   // hmiStns[3].wip[11].pnCode[4] := 1000;
   // hmiStns[3].wip[11].pnCode[5] := 1000;
   // hmiStns[3].wip[11].pnCode[6] := 1000;
   // hmiStns[3].wip[11].pnCode[7] := 1000;
   // hmiStns[3].wip[12].pnCode[0] := 1000;
   // hmiStns[3].wip[12].pnCode[1] := 1000;
   // hmiStns[3].wip[12].pnCode[2] := 1000;
   // hmiStns[3].wip[12].pnCode[3] := 1000;
   // hmiStns[3].wip[12].pnCode[4] := 1000;
   // hmiStns[3].wip[12].pnCode[5] := 1000;
   // hmiStns[3].wip[12].pnCode[6] := 1000;
   // hmiStns[3].wip[12].pnCode[7] := 1000;
   // hmiStns[3].wip[13].pnCode[0] := 1000;
   // hmiStns[3].wip[13].pnCode[1] := 1000;
   // hmiStns[3].wip[13].pnCode[2] := 1000;
   // hmiStns[3].wip[13].pnCode[3] := 1000;
   // hmiStns[3].wip[13].pnCode[4] := 1000;
   // hmiStns[3].wip[13].pnCode[5] := 1000;
   // hmiStns[3].wip[13].pnCode[6] := 1000;
   // hmiStns[3].wip[13].pnCode[7] := 1000;
   // hmiStns[3].wip[14].pnCode[0] := 1000;
   // hmiStns[3].wip[14].pnCode[1] := 1000;
   // hmiStns[3].wip[14].pnCode[2] := 1000;
   // hmiStns[3].wip[14].pnCode[3] := 1000;
   // hmiStns[3].wip[14].pnCode[4] := 1000;
   // hmiStns[3].wip[14].pnCode[5] := 1000;
   // hmiStns[3].wip[14].pnCode[6] := 1000;
   // hmiStns[3].wip[14].pnCode[7] := 1000;
   // hmiStns[3].wip[15].pnCode[0] := 1000;
   // hmiStns[3].wip[15].pnCode[1] := 1000;
   // hmiStns[3].wip[15].pnCode[2] := 1000;
   // hmiStns[3].wip[15].pnCode[3] := 1000;
   // hmiStns[3].wip[15].pnCode[4] := 1000;
   // hmiStns[3].wip[15].pnCode[5] := 1000;
   // hmiStns[3].wip[15].pnCode[6] := 1000;
   // hmiStns[3].wip[15].pnCode[7] := 1000;
   // hmiStns[3].wip[16].pnCode[0] := 1000;
   // hmiStns[3].wip[16].pnCode[1] := 1000;
   // hmiStns[3].wip[16].pnCode[2] := 1000;
   // hmiStns[3].wip[16].pnCode[3] := 1000;
   // hmiStns[3].wip[16].pnCode[4] := 1000;
   // hmiStns[3].wip[16].pnCode[5] := 1000;
   // hmiStns[3].wip[16].pnCode[6] := 1000;
   // hmiStns[3].wip[16].pnCode[7] := 1000;
   // hmiStns[3].wip[17].pnCode[0] := 1000;
   // hmiStns[3].wip[17].pnCode[1] := 1000;
   // hmiStns[3].wip[17].pnCode[2] := 1000;
   // hmiStns[3].wip[17].pnCode[3] := 1000;
   // hmiStns[3].wip[17].pnCode[4] := 1000;
   // hmiStns[3].wip[17].pnCode[5] := 1000;
   // hmiStns[3].wip[17].pnCode[6] := 1000;
   // hmiStns[3].wip[17].pnCode[7] := 1000;
   // hmiStns[3].wip[18].pnCode[0] := 1000;
   // hmiStns[3].wip[18].pnCode[1] := 1000;
   // hmiStns[3].wip[18].pnCode[2] := 1000;
   // hmiStns[3].wip[18].pnCode[3] := 1000;
   // hmiStns[3].wip[18].pnCode[4] := 1000;
   // hmiStns[3].wip[18].pnCode[5] := 1000;
   // hmiStns[3].wip[18].pnCode[6] := 1000;
   // hmiStns[3].wip[18].pnCode[7] := 1000;
   // hmiStns[3].wip[19].pnCode[0] := 1000;
   // hmiStns[3].wip[19].pnCode[1] := 1000;
   // hmiStns[3].wip[19].pnCode[2] := 1000;
   // hmiStns[3].wip[19].pnCode[3] := 1000;
   // hmiStns[3].wip[19].pnCode[4] := 1000;
   // hmiStns[3].wip[19].pnCode[5] := 1000;
   // hmiStns[3].wip[19].pnCode[6] := 1000;
   // hmiStns[3].wip[19].pnCode[7] := 1000;
   // hmiStns[3].wip[20].pnCode[0] := 1000;
   // hmiStns[3].wip[20].pnCode[1] := 1000;
   // hmiStns[3].wip[20].pnCode[2] := 1000;
   // hmiStns[3].wip[20].pnCode[3] := 1000;
   // hmiStns[3].wip[20].pnCode[4] := 1000;
   // hmiStns[3].wip[20].pnCode[5] := 1000;
   // hmiStns[3].wip[20].pnCode[6] := 1000;
   // hmiStns[3].wip[20].pnCode[7] := 1000;
   // hmiStns[3].wip[21].pnCode[0] := 1000;
   // hmiStns[3].wip[21].pnCode[1] := 1000;
   // hmiStns[3].wip[21].pnCode[2] := 1000;
   // hmiStns[3].wip[21].pnCode[3] := 1000;
   // hmiStns[3].wip[21].pnCode[4] := 1000;
   // hmiStns[3].wip[21].pnCode[5] := 1000;
   // hmiStns[3].wip[21].pnCode[6] := 1000;
   // hmiStns[3].wip[21].pnCode[7] := 1000;
   // hmiStns[3].wip[22].pnCode[0] := 1000;
   // hmiStns[3].wip[22].pnCode[1] := 1000;
   // hmiStns[3].wip[22].pnCode[2] := 1000;
   // hmiStns[3].wip[22].pnCode[3] := 1000;
   // hmiStns[3].wip[22].pnCode[4] := 1000;
   // hmiStns[3].wip[22].pnCode[5] := 1000;
   // hmiStns[3].wip[22].pnCode[6] := 1000;
   // hmiStns[3].wip[22].pnCode[7] := 1000;
   // hmiStns[3].wip[23].pnCode[0] := 1000;
   // hmiStns[3].wip[23].pnCode[1] := 1000;
   // hmiStns[3].wip[23].pnCode[2] := 1000;
   // hmiStns[3].wip[23].pnCode[3] := 1000;
   // hmiStns[3].wip[23].pnCode[4] := 1000;
   // hmiStns[3].wip[23].pnCode[5] := 1000;
   // hmiStns[3].wip[23].pnCode[6] := 1000;
   // hmiStns[3].wip[23].pnCode[7] := 1000;
   // hmiStns[3].wip[24].pnCode[0] := 1000;
   // hmiStns[3].wip[24].pnCode[1] := 1000;
   // hmiStns[3].wip[24].pnCode[2] := 1000;
   // hmiStns[3].wip[24].pnCode[3] := 1000;
   // hmiStns[3].wip[24].pnCode[4] := 1000;
   // hmiStns[3].wip[24].pnCode[5] := 1000;
   // hmiStns[3].wip[24].pnCode[6] := 1000;
   // hmiStns[3].wip[24].pnCode[7] := 1000;
   // hmiStns[3].wip[25].pnCode[0] := 1000;
   // hmiStns[3].wip[25].pnCode[1] := 1000;
   // hmiStns[3].wip[25].pnCode[2] := 1000;
   // hmiStns[3].wip[25].pnCode[3] := 1000;
   // hmiStns[3].wip[25].pnCode[4] := 1000;
   // hmiStns[3].wip[25].pnCode[5] := 1000;
   // hmiStns[3].wip[25].pnCode[6] := 1000;
   // hmiStns[3].wip[25].pnCode[7] := 1000;
   // hmiStns[3].wip[26].pnCode[0] := 1000;
   // hmiStns[3].wip[26].pnCode[1] := 1000;
   // hmiStns[3].wip[26].pnCode[2] := 1000;
   // hmiStns[3].wip[26].pnCode[3] := 1000;
   // hmiStns[3].wip[26].pnCode[4] := 1000;
   // hmiStns[3].wip[26].pnCode[5] := 1000;
   // hmiStns[3].wip[26].pnCode[6] := 1000;
   // hmiStns[3].wip[26].pnCode[7] := 1000;
   // hmiStns[3].wip[27].pnCode[0] := 1000;
   // hmiStns[3].wip[27].pnCode[1] := 1000;
   // hmiStns[3].wip[27].pnCode[2] := 1000;
   // hmiStns[3].wip[27].pnCode[3] := 1000;
   // hmiStns[3].wip[27].pnCode[4] := 1000;
   // hmiStns[3].wip[27].pnCode[5] := 1000;
   // hmiStns[3].wip[27].pnCode[6] := 1000;
   // hmiStns[3].wip[27].pnCode[7] := 1000;
   // hmiStns[3].wip[28].pnCode[0] := 1000;
   // hmiStns[3].wip[28].pnCode[1] := 1000;
   // hmiStns[3].wip[28].pnCode[2] := 1000;
   // hmiStns[3].wip[28].pnCode[3] := 1000;
   // hmiStns[3].wip[28].pnCode[4] := 1000;
   // hmiStns[3].wip[28].pnCode[5] := 1000;
   // hmiStns[3].wip[28].pnCode[6] := 1000;
   // hmiStns[3].wip[28].pnCode[7] := 1000;
   // hmiStns[3].wip[29].pnCode[0] := 1000;
   // hmiStns[3].wip[29].pnCode[1] := 1000;
   // hmiStns[3].wip[29].pnCode[2] := 1000;
   // hmiStns[3].wip[29].pnCode[3] := 1000;
   // hmiStns[3].wip[29].pnCode[4] := 1000;
   // hmiStns[3].wip[29].pnCode[5] := 1000;
   // hmiStns[3].wip[29].pnCode[6] := 1000;
   // hmiStns[3].wip[29].pnCode[7] := 1000;
   // hmiStns[3].wip[30].pnCode[0] := 1000;
   // hmiStns[3].wip[30].pnCode[1] := 1000;
   // hmiStns[3].wip[30].pnCode[2] := 1000;
   // hmiStns[3].wip[30].pnCode[3] := 1000;
   // hmiStns[3].wip[30].pnCode[4] := 1000;
   // hmiStns[3].wip[30].pnCode[5] := 1000;
   // hmiStns[3].wip[30].pnCode[6] := 1000;
   // hmiStns[3].wip[30].pnCode[7] := 1000;
   // hmiStns[3].wip[31].pnCode[0] := 1000;
   // hmiStns[3].wip[31].pnCode[1] := 1000;
   // hmiStns[3].wip[31].pnCode[2] := 1000;
   // hmiStns[3].wip[31].pnCode[3] := 1000;
   // hmiStns[3].wip[31].pnCode[4] := 1000;
   // hmiStns[3].wip[31].pnCode[5] := 1000;
   // hmiStns[3].wip[31].pnCode[6] := 1000;
   // hmiStns[3].wip[31].pnCode[7] := 1000;
   // hmiStns[3].wip[32].pnCode[0] := 1000;
   // hmiStns[3].wip[32].pnCode[1] := 1000;
   // hmiStns[3].wip[32].pnCode[2] := 1000;
   // hmiStns[3].wip[32].pnCode[3] := 1000;
   // hmiStns[3].wip[32].pnCode[4] := 1000;
   // hmiStns[3].wip[32].pnCode[5] := 1000;
   // hmiStns[3].wip[32].pnCode[6] := 1000;
   // hmiStns[3].wip[32].pnCode[7] := 1000;
   // hmiStns[3].wip[33].pnCode[0] := 1000;
   // hmiStns[3].wip[33].pnCode[1] := 1000;
   // hmiStns[3].wip[33].pnCode[2] := 1000;
   // hmiStns[3].wip[33].pnCode[3] := 1000;
   // hmiStns[3].wip[33].pnCode[4] := 1000;
   // hmiStns[3].wip[33].pnCode[5] := 1000;
   // hmiStns[3].wip[33].pnCode[6] := 1000;
   // hmiStns[3].wip[33].pnCode[7] := 1000;
   // hmiStns[3].wip[34].pnCode[0] := 1000;
   // hmiStns[3].wip[34].pnCode[1] := 1000;
   // hmiStns[3].wip[34].pnCode[2] := 1000;
   // hmiStns[3].wip[34].pnCode[3] := 1000;
   // hmiStns[3].wip[34].pnCode[4] := 1000;
   // hmiStns[3].wip[34].pnCode[5] := 1000;
   // hmiStns[3].wip[34].pnCode[6] := 1000;
   // hmiStns[3].wip[34].pnCode[7] := 1000;
   // hmiStns[3].wip[35].pnCode[0] := 1000;
   // hmiStns[3].wip[35].pnCode[1] := 1000;
   // hmiStns[3].wip[35].pnCode[2] := 1000;
   // hmiStns[3].wip[35].pnCode[3] := 1000;
   // hmiStns[3].wip[35].pnCode[4] := 1000;
   // hmiStns[3].wip[35].pnCode[5] := 1000;
   // hmiStns[3].wip[35].pnCode[6] := 1000;
   // hmiStns[3].wip[35].pnCode[7] := 1000;
   // hmiStns[3].wip[36].pnCode[0] := 1000;
   // hmiStns[3].wip[36].pnCode[1] := 1000;
   // hmiStns[3].wip[36].pnCode[2] := 1000;
   // hmiStns[3].wip[36].pnCode[3] := 1000;
   // hmiStns[3].wip[36].pnCode[4] := 1000;
   // hmiStns[3].wip[36].pnCode[5] := 1000;
   // hmiStns[3].wip[36].pnCode[6] := 1000;
   // hmiStns[3].wip[36].pnCode[7] := 1000;
   // hmiStns[3].wip[37].pnCode[0] := 1000;
   // hmiStns[3].wip[37].pnCode[1] := 1000;
   // hmiStns[3].wip[37].pnCode[2] := 1000;
   // hmiStns[3].wip[37].pnCode[3] := 1000;
   // hmiStns[3].wip[37].pnCode[4] := 1000;
   // hmiStns[3].wip[37].pnCode[5] := 1000;
   // hmiStns[3].wip[37].pnCode[6] := 1000;
   // hmiStns[3].wip[37].pnCode[7] := 1000;
   // hmiStns[3].wip[38].pnCode[0] := 1000;
   // hmiStns[3].wip[38].pnCode[1] := 1000;
   // hmiStns[3].wip[38].pnCode[2] := 1000;
   // hmiStns[3].wip[38].pnCode[3] := 1000;
   // hmiStns[3].wip[38].pnCode[4] := 1000;
   // hmiStns[3].wip[38].pnCode[5] := 1000;
   // hmiStns[3].wip[38].pnCode[6] := 1000;
   // hmiStns[3].wip[38].pnCode[7] := 1000;
   // hmiStns[3].wip[39].pnCode[0] := 1000;
   // hmiStns[3].wip[39].pnCode[1] := 1000;
   // hmiStns[3].wip[39].pnCode[2] := 1000;
   // hmiStns[3].wip[39].pnCode[3] := 1000;
   // hmiStns[3].wip[39].pnCode[4] := 1000;
   // hmiStns[3].wip[39].pnCode[5] := 1000;
   // hmiStns[3].wip[39].pnCode[6] := 1000;
   // hmiStns[3].wip[39].pnCode[7] := 1000;
   // hmiStns[3].wip[40].pnCode[0] := 1000;
   // hmiStns[3].wip[40].pnCode[1] := 1000;
   // hmiStns[3].wip[40].pnCode[2] := 1000;
   // hmiStns[3].wip[40].pnCode[3] := 1000;
   // hmiStns[3].wip[40].pnCode[4] := 1000;
   // hmiStns[3].wip[40].pnCode[5] := 1000;
   // hmiStns[3].wip[40].pnCode[6] := 1000;
   // hmiStns[3].wip[40].pnCode[7] := 1000;
   // hmiStns[3].wip[41].pnCode[0] := 1000;
   // hmiStns[3].wip[41].pnCode[1] := 1000;
   // hmiStns[3].wip[41].pnCode[2] := 1000;
   // hmiStns[3].wip[41].pnCode[3] := 1000;
   // hmiStns[3].wip[41].pnCode[4] := 1000;
   // hmiStns[3].wip[41].pnCode[5] := 1000;
   // hmiStns[3].wip[41].pnCode[6] := 1000;
   // hmiStns[3].wip[41].pnCode[7] := 1000;
   // hmiStns[3].wip[42].pnCode[0] := 1000;
   // hmiStns[3].wip[42].pnCode[1] := 1000;
   // hmiStns[3].wip[42].pnCode[2] := 1000;
   // hmiStns[3].wip[42].pnCode[3] := 1000;
   // hmiStns[3].wip[42].pnCode[4] := 1000;
   // hmiStns[3].wip[42].pnCode[5] := 1000;
   // hmiStns[3].wip[42].pnCode[6] := 1000;
   // hmiStns[3].wip[42].pnCode[7] := 1000;
   // hmiStns[3].wip[43].pnCode[0] := 1000;
   // hmiStns[3].wip[43].pnCode[1] := 1000;
   // hmiStns[3].wip[43].pnCode[2] := 1000;
   // hmiStns[3].wip[43].pnCode[3] := 1000;
   // hmiStns[3].wip[43].pnCode[4] := 1000;
   // hmiStns[3].wip[43].pnCode[5] := 1000;
   // hmiStns[3].wip[43].pnCode[6] := 1000;
   // hmiStns[3].wip[43].pnCode[7] := 1000;
   // hmiStns[3].wip[44].pnCode[0] := 1000;
   // hmiStns[3].wip[44].pnCode[1] := 1000;
   // hmiStns[3].wip[44].pnCode[2] := 1000;
   // hmiStns[3].wip[44].pnCode[3] := 1000;
   // hmiStns[3].wip[44].pnCode[4] := 1000;
   // hmiStns[3].wip[44].pnCode[5] := 1000;
   // hmiStns[3].wip[44].pnCode[6] := 1000;
   // hmiStns[3].wip[44].pnCode[7] := 1000;
   // hmiStns[3].wip[45].pnCode[0] := 1000;
   // hmiStns[3].wip[45].pnCode[1] := 1000;
   // hmiStns[3].wip[45].pnCode[2] := 1000;
   // hmiStns[3].wip[45].pnCode[3] := 1000;
   // hmiStns[3].wip[45].pnCode[4] := 1000;
   // hmiStns[3].wip[45].pnCode[5] := 1000;
   // hmiStns[3].wip[45].pnCode[6] := 1000;
   // hmiStns[3].wip[45].pnCode[7] := 1000;
   // hmiStns[3].wip[46].pnCode[0] := 1000;
   // hmiStns[3].wip[46].pnCode[1] := 1000;
   // hmiStns[3].wip[46].pnCode[2] := 1000;
   // hmiStns[3].wip[46].pnCode[3] := 1000;
   // hmiStns[3].wip[46].pnCode[4] := 1000;
   // hmiStns[3].wip[46].pnCode[5] := 1000;
   // hmiStns[3].wip[46].pnCode[6] := 1000;
   // hmiStns[3].wip[46].pnCode[7] := 1000;
   // hmiStns[3].wip[47].pnCode[0] := 1000;
   // hmiStns[3].wip[47].pnCode[1] := 1000;
   // hmiStns[3].wip[47].pnCode[2] := 1000;
   // hmiStns[3].wip[47].pnCode[3] := 1000;
   // hmiStns[3].wip[47].pnCode[4] := 1000;
   // hmiStns[3].wip[47].pnCode[5] := 1000;
   // hmiStns[3].wip[47].pnCode[6] := 1000;
   // hmiStns[3].wip[47].pnCode[7] := 1000;
   // hmiStns[3].wip[48].pnCode[0] := 1000;
   // hmiStns[3].wip[48].pnCode[1] := 1000;
   // hmiStns[3].wip[48].pnCode[2] := 1000;
   // hmiStns[3].wip[48].pnCode[3] := 1000;
   // hmiStns[3].wip[48].pnCode[4] := 1000;
   // hmiStns[3].wip[48].pnCode[5] := 1000;
   // hmiStns[3].wip[48].pnCode[6] := 1000;
   // hmiStns[3].wip[48].pnCode[7] := 1000;
   // hmiStns[3].wip[49].pnCode[0] := 1000;
   // hmiStns[3].wip[49].pnCode[1] := 1000;
   // hmiStns[3].wip[49].pnCode[2] := 1000;
   // hmiStns[3].wip[49].pnCode[3] := 1000;
   // hmiStns[3].wip[49].pnCode[4] := 1000;
   // hmiStns[3].wip[49].pnCode[5] := 1000;
   // hmiStns[3].wip[49].pnCode[6] := 1000;
   // hmiStns[3].wip[49].pnCode[7] := 1000;
   // hmiStns[4].pStn := 29;
   // hmiStns[4].wip[0].pnCode[0] := 1000;
   // hmiStns[4].wip[0].pnCode[1] := 244000;
   // hmiStns[4].wip[0].pnCode[2] := 1000;
   // hmiStns[4].wip[0].pnCode[3] := 4000;
   // hmiStns[4].wip[0].pnCode[4] := 1000;
   // hmiStns[4].wip[0].pnCode[5] := 1000;
   // hmiStns[4].wip[0].pnCode[6] := 2000;
   // hmiStns[4].wip[0].pnCode[7] := 3000;
   // hmiStns[4].wip[1].pnCode[0] := 1000;
   // hmiStns[4].wip[1].pnCode[1] := 244000;
   // hmiStns[4].wip[1].pnCode[2] := 6000;
   // hmiStns[4].wip[1].pnCode[3] := 10000;
   // hmiStns[4].wip[1].pnCode[4] := 1000;
   // hmiStns[4].wip[1].pnCode[5] := 7000;
   // hmiStns[4].wip[1].pnCode[6] := 5000;
   // hmiStns[4].wip[1].pnCode[7] := 11000;
   // hmiStns[4].wip[2].pnCode[0] := 1000;
   // hmiStns[4].wip[2].pnCode[1] := 244000;
   // hmiStns[4].wip[2].pnCode[2] := 8000;
   // hmiStns[4].wip[2].pnCode[3] := 10000;
   // hmiStns[4].wip[2].pnCode[4] := 1000;
   // hmiStns[4].wip[2].pnCode[5] := 9000;
   // hmiStns[4].wip[2].pnCode[6] := 5000;
   // hmiStns[4].wip[2].pnCode[7] := 11000;
   // hmiStns[4].wip[3].pnCode[0] := 1000;
   // hmiStns[4].wip[3].pnCode[1] := 1000;
   // hmiStns[4].wip[3].pnCode[2] := 1000;
   // hmiStns[4].wip[3].pnCode[3] := 1000;
   // hmiStns[4].wip[3].pnCode[4] := 1000;
   // hmiStns[4].wip[3].pnCode[5] := 1000;
   // hmiStns[4].wip[3].pnCode[6] := 1000;
   // hmiStns[4].wip[3].pnCode[7] := 1000;
   // hmiStns[4].wip[4].pnCode[0] := 1000;
   // hmiStns[4].wip[4].pnCode[1] := 1000;
   // hmiStns[4].wip[4].pnCode[2] := 1000;
   // hmiStns[4].wip[4].pnCode[3] := 1000;
   // hmiStns[4].wip[4].pnCode[4] := 1000;
   // hmiStns[4].wip[4].pnCode[5] := 1000;
   // hmiStns[4].wip[4].pnCode[6] := 1000;
   // hmiStns[4].wip[4].pnCode[7] := 1000;
   // hmiStns[4].wip[5].pnCode[0] := 1000;
   // hmiStns[4].wip[5].pnCode[1] := 1000;
   // hmiStns[4].wip[5].pnCode[2] := 1000;
   // hmiStns[4].wip[5].pnCode[3] := 1000;
   // hmiStns[4].wip[5].pnCode[4] := 1000;
   // hmiStns[4].wip[5].pnCode[5] := 1000;
   // hmiStns[4].wip[5].pnCode[6] := 1000;
   // hmiStns[4].wip[5].pnCode[7] := 1000;
   // hmiStns[4].wip[6].pnCode[0] := 1000;
   // hmiStns[4].wip[6].pnCode[1] := 1000;
   // hmiStns[4].wip[6].pnCode[2] := 1000;
   // hmiStns[4].wip[6].pnCode[3] := 1000;
   // hmiStns[4].wip[6].pnCode[4] := 1000;
   // hmiStns[4].wip[6].pnCode[5] := 1000;
   // hmiStns[4].wip[6].pnCode[6] := 1000;
   // hmiStns[4].wip[6].pnCode[7] := 1000;
   // hmiStns[4].wip[7].pnCode[0] := 1000;
   // hmiStns[4].wip[7].pnCode[1] := 1000;
   // hmiStns[4].wip[7].pnCode[2] := 1000;
   // hmiStns[4].wip[7].pnCode[3] := 1000;
   // hmiStns[4].wip[7].pnCode[4] := 1000;
   // hmiStns[4].wip[7].pnCode[5] := 1000;
   // hmiStns[4].wip[7].pnCode[6] := 1000;
   // hmiStns[4].wip[7].pnCode[7] := 1000;
   // hmiStns[4].wip[8].pnCode[0] := 1000;
   // hmiStns[4].wip[8].pnCode[1] := 1000;
   // hmiStns[4].wip[8].pnCode[2] := 1000;
   // hmiStns[4].wip[8].pnCode[3] := 1000;
   // hmiStns[4].wip[8].pnCode[4] := 1000;
   // hmiStns[4].wip[8].pnCode[5] := 1000;
   // hmiStns[4].wip[8].pnCode[6] := 1000;
   // hmiStns[4].wip[8].pnCode[7] := 1000;
   // hmiStns[4].wip[9].pnCode[0] := 1000;
   // hmiStns[4].wip[9].pnCode[1] := 1000;
   // hmiStns[4].wip[9].pnCode[2] := 1000;
   // hmiStns[4].wip[9].pnCode[3] := 1000;
   // hmiStns[4].wip[9].pnCode[4] := 1000;
   // hmiStns[4].wip[9].pnCode[5] := 1000;
   // hmiStns[4].wip[9].pnCode[6] := 1000;
   // hmiStns[4].wip[9].pnCode[7] := 1000;
   // hmiStns[4].wip[10].pnCode[0] := 1000;
   // hmiStns[4].wip[10].pnCode[1] := 1000;
   // hmiStns[4].wip[10].pnCode[2] := 1000;
   // hmiStns[4].wip[10].pnCode[3] := 1000;
   // hmiStns[4].wip[10].pnCode[4] := 1000;
   // hmiStns[4].wip[10].pnCode[5] := 1000;
   // hmiStns[4].wip[10].pnCode[6] := 1000;
   // hmiStns[4].wip[10].pnCode[7] := 1000;
   // hmiStns[4].wip[11].pnCode[0] := 1000;
   // hmiStns[4].wip[11].pnCode[1] := 1000;
   // hmiStns[4].wip[11].pnCode[2] := 1000;
   // hmiStns[4].wip[11].pnCode[3] := 1000;
   // hmiStns[4].wip[11].pnCode[4] := 1000;
   // hmiStns[4].wip[11].pnCode[5] := 1000;
   // hmiStns[4].wip[11].pnCode[6] := 1000;
   // hmiStns[4].wip[11].pnCode[7] := 1000;
   // hmiStns[4].wip[12].pnCode[0] := 1000;
   // hmiStns[4].wip[12].pnCode[1] := 1000;
   // hmiStns[4].wip[12].pnCode[2] := 1000;
   // hmiStns[4].wip[12].pnCode[3] := 1000;
   // hmiStns[4].wip[12].pnCode[4] := 1000;
   // hmiStns[4].wip[12].pnCode[5] := 1000;
   // hmiStns[4].wip[12].pnCode[6] := 1000;
   // hmiStns[4].wip[12].pnCode[7] := 1000;
   // hmiStns[4].wip[13].pnCode[0] := 1000;
   // hmiStns[4].wip[13].pnCode[1] := 1000;
   // hmiStns[4].wip[13].pnCode[2] := 1000;
   // hmiStns[4].wip[13].pnCode[3] := 1000;
   // hmiStns[4].wip[13].pnCode[4] := 1000;
   // hmiStns[4].wip[13].pnCode[5] := 1000;
   // hmiStns[4].wip[13].pnCode[6] := 1000;
   // hmiStns[4].wip[13].pnCode[7] := 1000;
   // hmiStns[4].wip[14].pnCode[0] := 1000;
   // hmiStns[4].wip[14].pnCode[1] := 1000;
   // hmiStns[4].wip[14].pnCode[2] := 1000;
   // hmiStns[4].wip[14].pnCode[3] := 1000;
   // hmiStns[4].wip[14].pnCode[4] := 1000;
   // hmiStns[4].wip[14].pnCode[5] := 1000;
   // hmiStns[4].wip[14].pnCode[6] := 1000;
   // hmiStns[4].wip[14].pnCode[7] := 1000;
   // hmiStns[4].wip[15].pnCode[0] := 1000;
   // hmiStns[4].wip[15].pnCode[1] := 1000;
   // hmiStns[4].wip[15].pnCode[2] := 1000;
   // hmiStns[4].wip[15].pnCode[3] := 1000;
   // hmiStns[4].wip[15].pnCode[4] := 1000;
   // hmiStns[4].wip[15].pnCode[5] := 1000;
   // hmiStns[4].wip[15].pnCode[6] := 1000;
   // hmiStns[4].wip[15].pnCode[7] := 1000;
   // hmiStns[4].wip[16].pnCode[0] := 1000;
   // hmiStns[4].wip[16].pnCode[1] := 1000;
   // hmiStns[4].wip[16].pnCode[2] := 1000;
   // hmiStns[4].wip[16].pnCode[3] := 1000;
   // hmiStns[4].wip[16].pnCode[4] := 1000;
   // hmiStns[4].wip[16].pnCode[5] := 1000;
   // hmiStns[4].wip[16].pnCode[6] := 1000;
   // hmiStns[4].wip[16].pnCode[7] := 1000;
   // hmiStns[4].wip[17].pnCode[0] := 1000;
   // hmiStns[4].wip[17].pnCode[1] := 1000;
   // hmiStns[4].wip[17].pnCode[2] := 1000;
   // hmiStns[4].wip[17].pnCode[3] := 1000;
   // hmiStns[4].wip[17].pnCode[4] := 1000;
   // hmiStns[4].wip[17].pnCode[5] := 1000;
   // hmiStns[4].wip[17].pnCode[6] := 1000;
   // hmiStns[4].wip[17].pnCode[7] := 1000;
   // hmiStns[4].wip[18].pnCode[0] := 1000;
   // hmiStns[4].wip[18].pnCode[1] := 1000;
   // hmiStns[4].wip[18].pnCode[2] := 1000;
   // hmiStns[4].wip[18].pnCode[3] := 1000;
   // hmiStns[4].wip[18].pnCode[4] := 1000;
   // hmiStns[4].wip[18].pnCode[5] := 1000;
   // hmiStns[4].wip[18].pnCode[6] := 1000;
   // hmiStns[4].wip[18].pnCode[7] := 1000;
   // hmiStns[4].wip[19].pnCode[0] := 1000;
   // hmiStns[4].wip[19].pnCode[1] := 1000;
   // hmiStns[4].wip[19].pnCode[2] := 1000;
   // hmiStns[4].wip[19].pnCode[3] := 1000;
   // hmiStns[4].wip[19].pnCode[4] := 1000;
   // hmiStns[4].wip[19].pnCode[5] := 1000;
   // hmiStns[4].wip[19].pnCode[6] := 1000;
   // hmiStns[4].wip[19].pnCode[7] := 1000;
   // hmiStns[4].wip[20].pnCode[0] := 1000;
   // hmiStns[4].wip[20].pnCode[1] := 1000;
   // hmiStns[4].wip[20].pnCode[2] := 1000;
   // hmiStns[4].wip[20].pnCode[3] := 1000;
   // hmiStns[4].wip[20].pnCode[4] := 1000;
   // hmiStns[4].wip[20].pnCode[5] := 1000;
   // hmiStns[4].wip[20].pnCode[6] := 1000;
   // hmiStns[4].wip[20].pnCode[7] := 1000;
   // hmiStns[4].wip[21].pnCode[0] := 1000;
   // hmiStns[4].wip[21].pnCode[1] := 1000;
   // hmiStns[4].wip[21].pnCode[2] := 1000;
   // hmiStns[4].wip[21].pnCode[3] := 1000;
   // hmiStns[4].wip[21].pnCode[4] := 1000;
   // hmiStns[4].wip[21].pnCode[5] := 1000;
   // hmiStns[4].wip[21].pnCode[6] := 1000;
   // hmiStns[4].wip[21].pnCode[7] := 1000;
   // hmiStns[4].wip[22].pnCode[0] := 1000;
   // hmiStns[4].wip[22].pnCode[1] := 1000;
   // hmiStns[4].wip[22].pnCode[2] := 1000;
   // hmiStns[4].wip[22].pnCode[3] := 1000;
   // hmiStns[4].wip[22].pnCode[4] := 1000;
   // hmiStns[4].wip[22].pnCode[5] := 1000;
   // hmiStns[4].wip[22].pnCode[6] := 1000;
   // hmiStns[4].wip[22].pnCode[7] := 1000;
   // hmiStns[4].wip[23].pnCode[0] := 1000;
   // hmiStns[4].wip[23].pnCode[1] := 1000;
   // hmiStns[4].wip[23].pnCode[2] := 1000;
   // hmiStns[4].wip[23].pnCode[3] := 1000;
   // hmiStns[4].wip[23].pnCode[4] := 1000;
   // hmiStns[4].wip[23].pnCode[5] := 1000;
   // hmiStns[4].wip[23].pnCode[6] := 1000;
   // hmiStns[4].wip[23].pnCode[7] := 1000;
   // hmiStns[4].wip[24].pnCode[0] := 1000;
   // hmiStns[4].wip[24].pnCode[1] := 1000;
   // hmiStns[4].wip[24].pnCode[2] := 1000;
   // hmiStns[4].wip[24].pnCode[3] := 1000;
   // hmiStns[4].wip[24].pnCode[4] := 1000;
   // hmiStns[4].wip[24].pnCode[5] := 1000;
   // hmiStns[4].wip[24].pnCode[6] := 1000;
   // hmiStns[4].wip[24].pnCode[7] := 1000;
   // hmiStns[4].wip[25].pnCode[0] := 1000;
   // hmiStns[4].wip[25].pnCode[1] := 1000;
   // hmiStns[4].wip[25].pnCode[2] := 1000;
   // hmiStns[4].wip[25].pnCode[3] := 1000;
   // hmiStns[4].wip[25].pnCode[4] := 1000;
   // hmiStns[4].wip[25].pnCode[5] := 1000;
   // hmiStns[4].wip[25].pnCode[6] := 1000;
   // hmiStns[4].wip[25].pnCode[7] := 1000;
   // hmiStns[4].wip[26].pnCode[0] := 1000;
   // hmiStns[4].wip[26].pnCode[1] := 1000;
   // hmiStns[4].wip[26].pnCode[2] := 1000;
   // hmiStns[4].wip[26].pnCode[3] := 1000;
   // hmiStns[4].wip[26].pnCode[4] := 1000;
   // hmiStns[4].wip[26].pnCode[5] := 1000;
   // hmiStns[4].wip[26].pnCode[6] := 1000;
   // hmiStns[4].wip[26].pnCode[7] := 1000;
   // hmiStns[4].wip[27].pnCode[0] := 1000;
   // hmiStns[4].wip[27].pnCode[1] := 1000;
   // hmiStns[4].wip[27].pnCode[2] := 1000;
   // hmiStns[4].wip[27].pnCode[3] := 1000;
   // hmiStns[4].wip[27].pnCode[4] := 1000;
   // hmiStns[4].wip[27].pnCode[5] := 1000;
   // hmiStns[4].wip[27].pnCode[6] := 1000;
   // hmiStns[4].wip[27].pnCode[7] := 1000;
   // hmiStns[4].wip[28].pnCode[0] := 1000;
   // hmiStns[4].wip[28].pnCode[1] := 1000;
   // hmiStns[4].wip[28].pnCode[2] := 1000;
   // hmiStns[4].wip[28].pnCode[3] := 1000;
   // hmiStns[4].wip[28].pnCode[4] := 1000;
   // hmiStns[4].wip[28].pnCode[5] := 1000;
   // hmiStns[4].wip[28].pnCode[6] := 1000;
   // hmiStns[4].wip[28].pnCode[7] := 1000;
   // hmiStns[4].wip[29].pnCode[0] := 1000;
   // hmiStns[4].wip[29].pnCode[1] := 1000;
   // hmiStns[4].wip[29].pnCode[2] := 1000;
   // hmiStns[4].wip[29].pnCode[3] := 1000;
   // hmiStns[4].wip[29].pnCode[4] := 1000;
   // hmiStns[4].wip[29].pnCode[5] := 1000;
   // hmiStns[4].wip[29].pnCode[6] := 1000;
   // hmiStns[4].wip[29].pnCode[7] := 1000;
   // hmiStns[4].wip[30].pnCode[0] := 1000;
   // hmiStns[4].wip[30].pnCode[1] := 1000;
   // hmiStns[4].wip[30].pnCode[2] := 1000;
   // hmiStns[4].wip[30].pnCode[3] := 1000;
   // hmiStns[4].wip[30].pnCode[4] := 1000;
   // hmiStns[4].wip[30].pnCode[5] := 1000;
   // hmiStns[4].wip[30].pnCode[6] := 1000;
   // hmiStns[4].wip[30].pnCode[7] := 1000;
   // hmiStns[4].wip[31].pnCode[0] := 1000;
   // hmiStns[4].wip[31].pnCode[1] := 1000;
   // hmiStns[4].wip[31].pnCode[2] := 1000;
   // hmiStns[4].wip[31].pnCode[3] := 1000;
   // hmiStns[4].wip[31].pnCode[4] := 1000;
   // hmiStns[4].wip[31].pnCode[5] := 1000;
   // hmiStns[4].wip[31].pnCode[6] := 1000;
   // hmiStns[4].wip[31].pnCode[7] := 1000;
   // hmiStns[4].wip[32].pnCode[0] := 1000;
   // hmiStns[4].wip[32].pnCode[1] := 1000;
   // hmiStns[4].wip[32].pnCode[2] := 1000;
   // hmiStns[4].wip[32].pnCode[3] := 1000;
   // hmiStns[4].wip[32].pnCode[4] := 1000;
   // hmiStns[4].wip[32].pnCode[5] := 1000;
   // hmiStns[4].wip[32].pnCode[6] := 1000;
   // hmiStns[4].wip[32].pnCode[7] := 1000;
   // hmiStns[4].wip[33].pnCode[0] := 1000;
   // hmiStns[4].wip[33].pnCode[1] := 1000;
   // hmiStns[4].wip[33].pnCode[2] := 1000;
   // hmiStns[4].wip[33].pnCode[3] := 1000;
   // hmiStns[4].wip[33].pnCode[4] := 1000;
   // hmiStns[4].wip[33].pnCode[5] := 1000;
   // hmiStns[4].wip[33].pnCode[6] := 1000;
   // hmiStns[4].wip[33].pnCode[7] := 1000;
   // hmiStns[4].wip[34].pnCode[0] := 1000;
   // hmiStns[4].wip[34].pnCode[1] := 1000;
   // hmiStns[4].wip[34].pnCode[2] := 1000;
   // hmiStns[4].wip[34].pnCode[3] := 1000;
   // hmiStns[4].wip[34].pnCode[4] := 1000;
   // hmiStns[4].wip[34].pnCode[5] := 1000;
   // hmiStns[4].wip[34].pnCode[6] := 1000;
   // hmiStns[4].wip[34].pnCode[7] := 1000;
   // hmiStns[4].wip[35].pnCode[0] := 1000;
   // hmiStns[4].wip[35].pnCode[1] := 1000;
   // hmiStns[4].wip[35].pnCode[2] := 1000;
   // hmiStns[4].wip[35].pnCode[3] := 1000;
   // hmiStns[4].wip[35].pnCode[4] := 1000;
   // hmiStns[4].wip[35].pnCode[5] := 1000;
   // hmiStns[4].wip[35].pnCode[6] := 1000;
   // hmiStns[4].wip[35].pnCode[7] := 1000;
   // hmiStns[4].wip[36].pnCode[0] := 1000;
   // hmiStns[4].wip[36].pnCode[1] := 1000;
   // hmiStns[4].wip[36].pnCode[2] := 1000;
   // hmiStns[4].wip[36].pnCode[3] := 1000;
   // hmiStns[4].wip[36].pnCode[4] := 1000;
   // hmiStns[4].wip[36].pnCode[5] := 1000;
   // hmiStns[4].wip[36].pnCode[6] := 1000;
   // hmiStns[4].wip[36].pnCode[7] := 1000;
   // hmiStns[4].wip[37].pnCode[0] := 1000;
   // hmiStns[4].wip[37].pnCode[1] := 1000;
   // hmiStns[4].wip[37].pnCode[2] := 1000;
   // hmiStns[4].wip[37].pnCode[3] := 1000;
   // hmiStns[4].wip[37].pnCode[4] := 1000;
   // hmiStns[4].wip[37].pnCode[5] := 1000;
   // hmiStns[4].wip[37].pnCode[6] := 1000;
   // hmiStns[4].wip[37].pnCode[7] := 1000;
   // hmiStns[4].wip[38].pnCode[0] := 1000;
   // hmiStns[4].wip[38].pnCode[1] := 1000;
   // hmiStns[4].wip[38].pnCode[2] := 1000;
   // hmiStns[4].wip[38].pnCode[3] := 1000;
   // hmiStns[4].wip[38].pnCode[4] := 1000;
   // hmiStns[4].wip[38].pnCode[5] := 1000;
   // hmiStns[4].wip[38].pnCode[6] := 1000;
   // hmiStns[4].wip[38].pnCode[7] := 1000;
   // hmiStns[4].wip[39].pnCode[0] := 1000;
   // hmiStns[4].wip[39].pnCode[1] := 1000;
   // hmiStns[4].wip[39].pnCode[2] := 1000;
   // hmiStns[4].wip[39].pnCode[3] := 1000;
   // hmiStns[4].wip[39].pnCode[4] := 1000;
   // hmiStns[4].wip[39].pnCode[5] := 1000;
   // hmiStns[4].wip[39].pnCode[6] := 1000;
   // hmiStns[4].wip[39].pnCode[7] := 1000;
   // hmiStns[4].wip[40].pnCode[0] := 1000;
   // hmiStns[4].wip[40].pnCode[1] := 1000;
   // hmiStns[4].wip[40].pnCode[2] := 1000;
   // hmiStns[4].wip[40].pnCode[3] := 1000;
   // hmiStns[4].wip[40].pnCode[4] := 1000;
   // hmiStns[4].wip[40].pnCode[5] := 1000;
   // hmiStns[4].wip[40].pnCode[6] := 1000;
   // hmiStns[4].wip[40].pnCode[7] := 1000;
   // hmiStns[4].wip[41].pnCode[0] := 1000;
   // hmiStns[4].wip[41].pnCode[1] := 1000;
   // hmiStns[4].wip[41].pnCode[2] := 1000;
   // hmiStns[4].wip[41].pnCode[3] := 1000;
   // hmiStns[4].wip[41].pnCode[4] := 1000;
   // hmiStns[4].wip[41].pnCode[5] := 1000;
   // hmiStns[4].wip[41].pnCode[6] := 1000;
   // hmiStns[4].wip[41].pnCode[7] := 1000;
   // hmiStns[4].wip[42].pnCode[0] := 1000;
   // hmiStns[4].wip[42].pnCode[1] := 1000;
   // hmiStns[4].wip[42].pnCode[2] := 1000;
   // hmiStns[4].wip[42].pnCode[3] := 1000;
   // hmiStns[4].wip[42].pnCode[4] := 1000;
   // hmiStns[4].wip[42].pnCode[5] := 1000;
   // hmiStns[4].wip[42].pnCode[6] := 1000;
   // hmiStns[4].wip[42].pnCode[7] := 1000;
   // hmiStns[4].wip[43].pnCode[0] := 1000;
   // hmiStns[4].wip[43].pnCode[1] := 1000;
   // hmiStns[4].wip[43].pnCode[2] := 1000;
   // hmiStns[4].wip[43].pnCode[3] := 1000;
   // hmiStns[4].wip[43].pnCode[4] := 1000;
   // hmiStns[4].wip[43].pnCode[5] := 1000;
   // hmiStns[4].wip[43].pnCode[6] := 1000;
   // hmiStns[4].wip[43].pnCode[7] := 1000;
   // hmiStns[4].wip[44].pnCode[0] := 1000;
   // hmiStns[4].wip[44].pnCode[1] := 1000;
   // hmiStns[4].wip[44].pnCode[2] := 1000;
   // hmiStns[4].wip[44].pnCode[3] := 1000;
   // hmiStns[4].wip[44].pnCode[4] := 1000;
   // hmiStns[4].wip[44].pnCode[5] := 1000;
   // hmiStns[4].wip[44].pnCode[6] := 1000;
   // hmiStns[4].wip[44].pnCode[7] := 1000;
   // hmiStns[4].wip[45].pnCode[0] := 1000;
   // hmiStns[4].wip[45].pnCode[1] := 1000;
   // hmiStns[4].wip[45].pnCode[2] := 1000;
   // hmiStns[4].wip[45].pnCode[3] := 1000;
   // hmiStns[4].wip[45].pnCode[4] := 1000;
   // hmiStns[4].wip[45].pnCode[5] := 1000;
   // hmiStns[4].wip[45].pnCode[6] := 1000;
   // hmiStns[4].wip[45].pnCode[7] := 1000;
   // hmiStns[4].wip[46].pnCode[0] := 1000;
   // hmiStns[4].wip[46].pnCode[1] := 1000;
   // hmiStns[4].wip[46].pnCode[2] := 1000;
   // hmiStns[4].wip[46].pnCode[3] := 1000;
   // hmiStns[4].wip[46].pnCode[4] := 1000;
   // hmiStns[4].wip[46].pnCode[5] := 1000;
   // hmiStns[4].wip[46].pnCode[6] := 1000;
   // hmiStns[4].wip[46].pnCode[7] := 1000;
   // hmiStns[4].wip[47].pnCode[0] := 1000;
   // hmiStns[4].wip[47].pnCode[1] := 1000;
   // hmiStns[4].wip[47].pnCode[2] := 1000;
   // hmiStns[4].wip[47].pnCode[3] := 1000;
   // hmiStns[4].wip[47].pnCode[4] := 1000;
   // hmiStns[4].wip[47].pnCode[5] := 1000;
   // hmiStns[4].wip[47].pnCode[6] := 1000;
   // hmiStns[4].wip[47].pnCode[7] := 1000;
   // hmiStns[4].wip[48].pnCode[0] := 1000;
   // hmiStns[4].wip[48].pnCode[1] := 1000;
   // hmiStns[4].wip[48].pnCode[2] := 1000;
   // hmiStns[4].wip[48].pnCode[3] := 1000;
   // hmiStns[4].wip[48].pnCode[4] := 1000;
   // hmiStns[4].wip[48].pnCode[5] := 1000;
   // hmiStns[4].wip[48].pnCode[6] := 1000;
   // hmiStns[4].wip[48].pnCode[7] := 1000;
   // hmiStns[4].wip[49].pnCode[0] := 1000;
   // hmiStns[4].wip[49].pnCode[1] := 1000;
   // hmiStns[4].wip[49].pnCode[2] := 1000;
   // hmiStns[4].wip[49].pnCode[3] := 1000;
   // hmiStns[4].wip[49].pnCode[4] := 1000;
   // hmiStns[4].wip[49].pnCode[5] := 1000;
   // hmiStns[4].wip[49].pnCode[6] := 1000;
   // hmiStns[4].wip[49].pnCode[7] := 1000;
   // // kp8Stns[0] : VOLVO 16 01
   // // kp8Stns[1] : VOLVO 16 02
   // // kp8Stns[2] : VOLVO 16 03
   // // kp8Stns[3] : VOLVO 16 04
   // // kp8Stns[4] : VOLVO 16 05
   // // kp8Stns[5] : VOLVO 16 06
   // // kp8Stns[6] : VOLVO 16 07
   // // kp8Stns[7] : VOLVO 16 08
   // // kp8Stns[8] : VOLVO 16 09
   // // kp8Stns[9] : VOLVO 16 10
   // // kp8Stns[10] : VOLVO 16 11
   // // kp8Stns[11] : CHM 01
   // // kp8Stns[12] : CHM 02
   // // kp8Stns[13] : CHM 03
   // // kp8Stns[14] : CHM 04
   // // kp8Stns[15] : CHM 05
   // // kp8Stns[16] : CDO 01
   // // kp8Stns[17] : CDO 02
   // // kp8Stns[18] : CDO 03
   // // kp8Stns[19] : BFL 01
   // // kp8Stns[20] : BFL 02
   // // kp8Stns[21] : BFL 03
   // // kp8Stns[22] : LGS 01
   // // kp8Stns[23] : LGS 02
   // // kp8Stns[24] : LGS 03
   // // kp8Stns[25] : PC 02
   // // kp8Stns[26] : 1BX2.0 01
   // // kp8Stns[27] : 1BX2.0 02
   // // kp8Stns[28] : 1BX2.0 03
   // // kp8Stns[29] : 1BX2.0 04
   // // kp8Stns[30] : 1BX2.0 05
   // // kp8Stns[31] : 1BX3.0 01
   // // kp8Stns[32] : 1BX3.0 02
   // // kp8Stns[33] : 1BX3.0 03
   // // hmiStns[0] : CV 01
   // // hmiStns[1] : CV 02
   // // hmiStns[2] : CV 03
   // // hmiStns[3] : CV 04
   // // hmiStns[4] : PC 01
END_TYPE

// folder: HMI Station

TYPE "HMI Station: Part Selection Screen"
   STRUCT
      animate : Array[0.."partSelScrnObjCnt"] of Int;
      pbs : DWord;
      txt : Array[0.."partSelScrnObjCnt"] of WString [40];
   END_STRUCT;
END_TYPE

TYPE "HMI Stations"
   STRUCT
      stns : Array[0.."hmi_station_count"] of "HMI Station: Compressed";
   END_STRUCT;
END_TYPE

TYPE "HMI Station: Wip Select: PLC Interface"
   STRUCT
      raw : Array[0..31] of Bool;
      wsRising : Array[0..5] of Bool;
      wsFalling : Array[0..5] of Bool;
   END_STRUCT;
END_TYPE

TYPE "HMI Station: Compressed"
   STRUCT
      partSelect : "HMI Station: Part Selection Screen";
      template : "HMI Station: Template Screen";
      wipSelect : "HMI Station: Wip Select: Screen";
   END_STRUCT;
END_TYPE

